(* Logix 5000 project; controller _GigaDiscovery vendor 1 type 14 code 244 rev 35.11; software revision 35.03; part 5 of 23 *)
(* tags used below, declared in another part *)
   All_RESTRAINTS_Opened : BOOL;
   Analog_Input_Pos_6 : REAL[8];
   Compressor_Pressure_OK : BOOL;
   Emergencies_CL1 : DINT[14];
   Gates_Open_Permissive : Permissive;
   Girella_Field_Actuate_During_Inactivity : BOOL;
   Girella_Gradi_Sec : DINT;
   Gondola_Axe : Axe;
   HMI_Light_Pb : BOOL;
   HMI_Status_Safety : Status_Safety;
   I_ADSL_Fault_Ch1 : BOOL;   // Gondola Communication Modem Fault CH1 -T27002C
   I_ADSL_Fault_Ch2 : BOOL;   // Gondola Communication Modem Fault CH2 -T27002C
   I_Compressor_Motor_Protection : BOOL;   // Compressor Motor Protection Feedback -F18002C
   I_Dryer_Motor_Protection : BOOL;   // Dryer Motor Protection Feedback -F18202C
   I_Gate_1_Opened : BOOL;   // Gate 1 RFID Sensor Closed -B24501J
   I_Gate_2_Opened : BOOL;   // Gate 2 RFID Sensor Closed -B24601J
   I_Gate_3_Opened : BOOL;   // Gate 3 RFID Sensor Closed -B24701J
   I_Gate_4_Opened : BOOL;   // Gate 4 RFID Sensor Closed -B24801J
   I_Light_Selector : BOOL;   // Light Selector Switch -S30408F
   I_Motor_1_2_Fan_Protection_Feedback : BOOL;   // Motor 1-2 Fan Protection Feedback -F10402C -F10406C
   I_Motor_1_Overvoltage_Control : BOOL;   // Motor 1 Overvoltage control - Relay OK -K10302G
   I_Motor_1_Thermal_Probe : BOOL;   // Motor 1 Thermal Probe -K10702H
   I_Motor_2_Overvoltage_Control : BOOL;   // Motor 2 Overvoltage control - Relay OK -K10307G
   I_Motor_2_Thermal_Probe : BOOL;   // Motor 2 Thermal Probe -K10704H
   I_Motor_3_4_Fan_Protection_Feedback : BOOL;   // Motor 3-4 Fan Protection Feedback -F12402C -F12406C
   I_Motor_3_Overvoltage_Control : BOOL;   // Motor 3 Overvoltage control - Relay OK -K12302G
   I_Motor_3_Thermal_Probe : BOOL;   // Motor 3 Thermal Probe -K12702H
   I_Motor_4_Overvoltage_Control : BOOL;   // Motor 4 Overvoltage control - Relay OK -K12307G
   I_Motor_4_Thermal_Probe : BOOL;   // Motor 4 Thermal Probe -K12704H
   I_Motor_5_6_Fan_Protection_Feedback : BOOL;   // Motor 5-6 Fan Protection Feedback -F14402C -F14406C
   I_Motor_5_Overvoltage_Control : BOOL;   // Motor 5 Overvoltage control - Relay OK -K14302G
   I_Motor_5_Thermal_Probe : BOOL;   // Motor 5 Thermal Probe -K14702H
   I_Motor_6_Overvoltage_Control : BOOL;   // Motor 6 Overvoltage control - Relay OK -K14307G
   I_Motor_6_Thermal_Probe : BOOL;   // Motor 6 Thermal Probe -K14704H
   I_Motor_7_Fan_Protection_Feedback : BOOL;   // Motor 7 Fan Protection Feedback -F16402C
   I_Motor_7_Thermal_Probe : BOOL;   // Motor 7 Thermal Probe -K16602H
   I_OCC_Operator_Enable_Key : BOOL;   // OCC Console Enabled -S30305F
   I_Platform_Closed : UDT_DCM;   // Platform Closed RFID Series -B22501J... -B22807J -B22801B
   I_Platform_Opened : UDT_DCM;   // Platform Opened RFID Series -Q23801J -Q23807J
   I_Remote_Connection_Enabled : BOOL;   // Remote Connection active ROUTER eWON K74A04E
   K_Speed : REAL;
   MCC_71_03 : BOOL[32];
   MODE : BOOL;   // MODE 0 = AUTO 1 = MANUAL -S30801F
   NO_SFTY_GateClosedSeries : BOOL;   // All Gates Closed and Locked
   O_Close_Gates : BOOL;
   ONP : DINT;   // Optional Not Present
   Pb_Platform_Stop : BOOL;   // Platform Stop Command -S30608F
   Platform_Close_Cycle : Sequencer;
   Platform_Close_Permissive : Permissive;
   Platform_Open_Cycle : Sequencer;
   Platform_Open_Permissive : Permissive;
   Pylon_Axe : Axe;
   Pylon_Field_Actuate_During_Inactivity : BOOL;
   Real : REAL[32];
   RESTRAINTS_Closed : BOOL;   // All RESTRAINTS Closed
   Restraints_Cycle : Sequencer;
   Restraints_Permissive : Permissive;
   Start_Permissive : Permissive;
   Start_Permissive2 : Permissive;
   Start_Stop_Cycle : Sequencer;
   Test : DCI_STOP_TEST;
   To_Sfty : Std_to_Sfty;
(* General, continued *)

ROUTINE Main   (* ladder *)
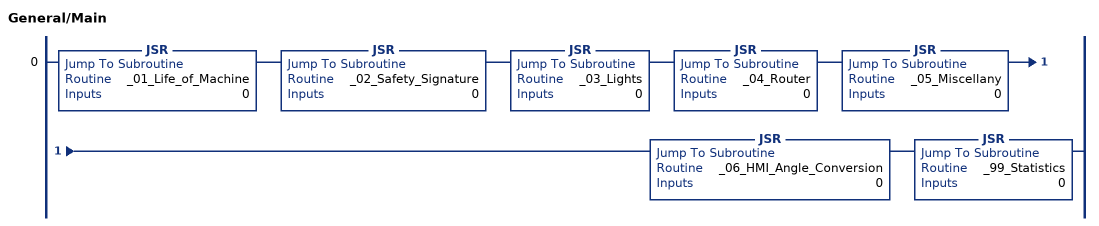
   0: JSR(_01_Life_of_Machine,0)JSR(_02_Safety_Signature,0)JSR(_03_Lights,0)JSR(_04_Router,0)JSR(_05_Miscellany,0)JSR(_06_HMI_Angle_Conversion,0)JSR(_99_Statistics,0);
END_ROUTINE
END_PROGRAM

PROGRAM HMI   (* main routine Main *)
VAR
   HMI_Auto_Cycle_Permissive : Permissive_Description := (Visible_Bits := 2147475455, Header_Description_en := 'Start Permissives (1)', Header_Description_others := 'Permessi di Start (1)', Bit_Description_en[0] := 'OCC2 Allow Main Confirm -S28602F', Bit_Description_en[1] := 'OCC Console Enabled -S30305F', Bit_Description_en[2] := 'OCC Stop Button Not Pressed -S30308F', Bit_Description_en[3] := 'All Restraints Closed', Bit_Description_en[4] := 'Gates 01-04 Closed -B24602J....-B24802J', Bit_Description_en[5] := 'Platform Stop Command Not Pressed -S30608F', Bit_Description_en[6] := 'No Emergencies Class 0', Bit_Description_en[7] := 'Restraints Proof Test Ok', Bit_Description_en[8] := 'OCC Motion Lockout -Q31203E', Bit_Description_en[9] := 'Restraints Main Valve Limit Switch Closed -B40508I', Bit_Description_en[10] := 'OCC2 E-Stop PB Not Pressed -S28502F', Bit_Description_en[11] := 'Platform Main Valve Closed -B21902I', Bit_Description_en[12] := 'Pylon Minimum Speed', Bit_Description_en[13] := 'Restraints Main Valve Pressure Switch Closed -S40602J', Bit_Description_en[14] := 'Power On Delay (80 sec.)', Bit_Description_en[15] := 'Restraints Opened Correctly', Bit_Description_en[16] := 'Restraints Pressure Switches Working Correctly', Bit_Description_en[17] := 'No Emergencies Class 1', Bit_Description_en[18] := 'Restraints Closed Correctly', Bit_Description_en[19] := 'OCC Footpedal Memory -S30901F', Bit_Description_en[20] := 'Valves Proof Test OK', Bit_Description_en[21] := 'Pylon Motors Fan On -Q9302F', Bit_Description_en[22] := 'OCC E-Stop PB Test Ok -S30301F', Bit_Description_en[23] := 'Motor Field Contactors All Disabled -Q10101E -Q10103E -Q16105E -Q16107E', Bit_Description_en[24] := 'Pylon Stopped at Home Position -B26002I -B26007I', Bit_Description_en[25] := 'Line Minimum Pressure -S21504B', Bit_Description_en[26] := 'Restraints Racks Unlock Valve Pressure Ok', Bit_Description_en[27] := 'All Racks Closed', Bit_Description_en[28] := 'Platform Opened -Q28301J -Q23807J', Bit_Description_en[29] := 'Gate Exit (G05) Closed -B25304I', Bit_Description_en[30] := 'Gate Enter (G01) Closed -B25204I', Bit_Description_en[31] := 'Gate 4 Operator(MOP) Closed -B25404J');
   HMI_Auto_Cycle_Permissive2 : Permissive_Description := (Visible_Bits := 255, Header_Description_en := 'Start Permissives (2)', Header_Description_others := 'Permessi di Start (2)', Bit_Description_en[0] := 'Platform Line Minimum Pressure Switch Closed -S21511B', Bit_Description_en[1] := 'Platform Pilot Valves Not Enabled to Open/Close -Y22002A', Bit_Description_en[2] := 'Restraints Main Valve Limit Switch Closed -B5408I', Bit_Description_en[3] := 'Restraints Sectors Left and Right Valves Unlock Disabled', Bit_Description_en[4] := 'All Restraints Sectors Disabled', Bit_Description_en[5] := 'OCC2 Stop PB Not Pressed -S28606F', Bit_Description_en[6] := 'Main Valve Closed -B40501I', Bit_Description_en[7] := 'All Restraints Sectors Racks On');
   HMI_Gates_Open_Permissive : Permissive_Description := (FailBitsConditions := 16, Visible_Bits := 190, Header_Description_en := 'Gates Open Permissives', Header_Description_others := 'Permessi di Apertura dei Cancelli', Bit_Description_en[1] := 'Ride Not in Start', Bit_Description_en[2] := 'Gondola Minimum Speed', Bit_Description_en[3] := 'Platform Main Valve Not Commanded -B21920I', Bit_Description_en[4] := 'Platform Closed -B22501J...-B22807J -B22801B', Bit_Description_en[5] := 'Pylon Safety Angle', Bit_Description_en[7] := 'Pylon Minimum Speed');
   HMI_Night_Mode : BOOL;
   HMI_Platform_Close_Error : BOOL;
   HMI_Platform_Close_Permissive : Permissive_Description := (OS_Fail := 1, Visible_Bits := 16375, Header_Description_en := 'Platform Close Permissives', Header_Description_others := 'Permessi di Chiusura della Piattaforma', Bit_Description_en[0] := 'OCC E-Stop PB Not Pressed -S30301F', Bit_Description_en[1] := 'Power On Delay (80 sec.)', Bit_Description_en[2] := 'OCC Console Enabled -S30305F', Bit_Description_en[4] := 'Motor Field Contactors All Disabled -Q10101E -Q10103E -Q16105E -Q16107E', Bit_Description_en[5] := 'Pylon Stoped At Home Position -B26002I -B26007I', Bit_Description_en[6] := 'Compressor Minimum Pressure -S21504B', Bit_Description_en[7] := 'Platform Close Alarms Not Present', Bit_Description_en[8] := 'Pylon Safety Angle', Bit_Description_en[9] := 'Pylon Minimum Speed', Bit_Description_en[10] := 'Gondola Minimun Speed', Bit_Description_en[11] := 'Platform Stop Push Button Not Pressed -S30608F', Bit_Description_en[12] := 'OCC Motion Lockout -Q31203E', Bit_Description_en[13] := 'OCC2 E-Stop PB Not Pressed -S28502F');
   HMI_Platform_Closed : BOOL := 1;
   HMI_Platform_Closing : BOOL;
   HMI_Platform_Open_Error : BOOL;
   HMI_Platform_Open_Permissive : Permissive_Description := (Visible_Bits := -2097153, Header_Description_en := 'Platform Open Permissives', Header_Description_others := 'Permessi di Apertura della Piattaforma', Bit_Description_en[0] := 'OCC E-Stop PB Not Pressed -S30301F', Bit_Description_en[1] := 'Power On Delay (80 sec.)', Bit_Description_en[2] := 'OCC Console Enabled -S3201E', Bit_Description_en[3] := 'Restraints Closed', Bit_Description_en[4] := 'Main Valve Closed -B40501I', Bit_Description_en[5] := 'Ride Not in Start', Bit_Description_en[6] := 'Compressor Minimum Pressure ', Bit_Description_en[7] := 'OCC Stop Button Not Pressed -S30308F', Bit_Description_en[8] := 'Gates 01-04 Closed -B24602J....-B24802J', Bit_Description_en[9] := 'Platform Stop Push Button not Pressed -S30608F', Bit_Description_en[10] := 'No Emergencies', Bit_Description_en[11] := 'OCC2 Allow Main Confirm -S28602F', Bit_Description_en[12] := 'OCC2 E-Stop PB Not Pressed -S28502F', Bit_Description_en[13] := 'OCC Motion Lockout -Q31203E', Bit_Description_en[14] := 'All Restraints Sectors Disabled', Bit_Description_en[15] := 'Gate Exit (G05) Closed -B25304I', Bit_Description_en[16] := 'Gate Enter (G01) Closed -B25204I', Bit_Description_en[17] := 'Gate 4 Operator(MOP) Closed -B25404J', Bit_Description_en[18] := 'Restraints Proof Test Ok', Bit_Description_en[19] := 'Restraints Main Valve Limit Switch Closed -B40508I', Bit_Description_en[20] := 'Pylon Minimum Speed', Bit_Description_en[22] := 'Restraints Opened Correctly', Bit_Description_en[23] := 'Restraints Pressure Switches Working Correctly', Bit_Description_en[24] := 'Restraints Closed Correctly', Bit_Description_en[25] := 'OCC Footpedal Memory -S30901F', Bit_Description_en[26] := 'Pylon Motors Fan On -Q9302F', Bit_Description_en[27] := 'Motor Field Contactors All Disabled -Q10101E -Q10103E -Q16105E -Q16107E', Bit_Description_en[28] := 'Pylon Stopped at Home Position -B26002I -B26007I', Bit_Description_en[29] := 'All Racks Closed', Bit_Description_en[30] := 'OCC2 Stop PB Not Pressed -S28606F', Bit_Description_en[31] := 'Platform Not at Maximum Closing Pressure -S21510B');
   HMI_Platform_Opened : BOOL;
   HMI_Platform_Opening : BOOL;
   HMI_Restraints_Closed : BOOL := 1;
   HMI_Restraints_Closing : BOOL;
   HMI_Restraints_Error : BOOL;
   HMI_Restraints_Opened : BOOL;
   HMI_Restraints_Opening : BOOL;
   HMI_Restraints_Permissive : Permissive_Description := (Visible_Bits := 7274495, Header_Description_en := 'Restraints Release Permissives', Header_Description_others := 'Permessi di Rilascio dei Maniglioni', Bit_Description_en[0] := 'OCC E-Stop PB Not Pressed -S30301F', Bit_Description_en[1] := 'Power On Delay (80 sec.)', Bit_Description_en[2] := 'OCC Console Enabled -S30305F', Bit_Description_en[3] := 'Platform Closed Cycle Complete', Bit_Description_en[4] := 'Platform Not at Maximum Closing Pressure -S21510B', Bit_Description_en[5] := 'Ride Not in Start', Bit_Description_en[6] := 'Pylon Stopped at Home Position -B26002I -B26007I', Bit_Description_en[7] := 'Pylon Encoder Low Position', Bit_Description_en[8] := 'Pylon Low Speed', Bit_Description_en[9] := 'Gondola Low Speed', Bit_Description_en[10] := 'All Pylon and Gondola Drives Not Running', Bit_Description_en[11] := 'Motor Field Contactors All Disabled -Q10101E -Q10103E -Q16105E -Q16107E', Bit_Description_en[12] := 'OCC2 E-Stop PB Not Pressed -S28502F', Bit_Description_en[13] := 'OCC Motion Lockout -Q31203E', Bit_Description_en[14] := 'Retraints Not Opened During ProofTest', Bit_Description_en[15] := 'Platform Main Valve Open -B21902I', Bit_Description_en[17] := 'Platform Line Minimum Pressure Switch Closed -S21511B', Bit_Description_en[18] := 'Platform Pilot Valves Not Enabled to Open/Close -Y22002A', Bit_Description_en[19] := 'Unlock Platform Line Pressure Switch Open -S22006B', Bit_Description_en[21] := 'Platform Closed', Bit_Description_en[22] := 'Platform Not Open');
   Os : SINT := 20;
END_VAR

ROUTINE HMI_Permissive   (* ladder *)
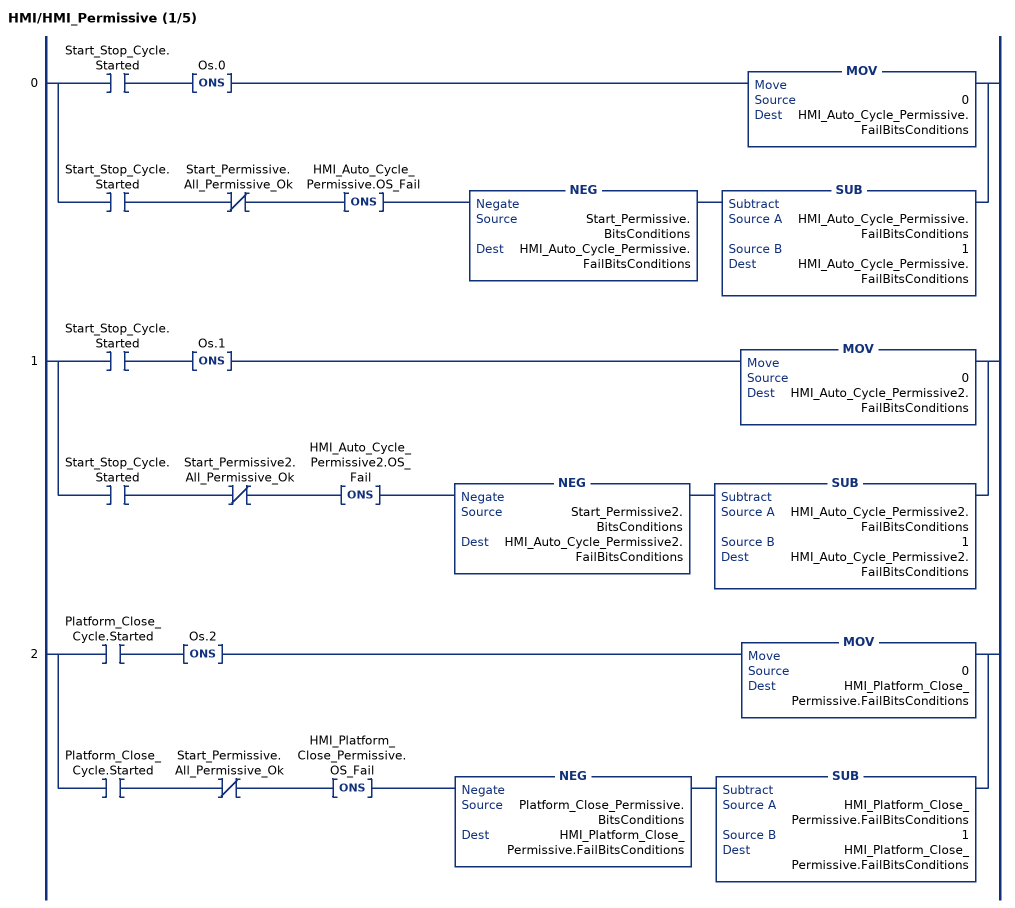
   0: [XIC(Start_Stop_Cycle.Started) ONS(Os.0) MOV(0,HMI_Auto_Cycle_Permissive.FailBitsConditions) ,XIC(Start_Stop_Cycle.Started) XIO(Start_Permissive.All_Permissive_Ok) ONS(HMI_Auto_Cycle_Permissive.OS_Fail) NEG(Start_Permissive.BitsConditions,HMI_Auto_Cycle_Permissive.FailBitsConditions) SUB(HMI_Auto_Cycle_Permissive.FailBitsConditions,1,HMI_Auto_Cycle_Permissive.FailBitsConditions) ];
   1: [XIC(Start_Stop_Cycle.Started) ONS(Os.1) MOV(0,HMI_Auto_Cycle_Permissive2.FailBitsConditions) ,XIC(Start_Stop_Cycle.Started) XIO(Start_Permissive2.All_Permissive_Ok) ONS(HMI_Auto_Cycle_Permissive2.OS_Fail) NEG(Start_Permissive2.BitsConditions,HMI_Auto_Cycle_Permissive2.FailBitsConditions) SUB(HMI_Auto_Cycle_Permissive2.FailBitsConditions,1,HMI_Auto_Cycle_Permissive2.FailBitsConditions) ];
   2: [XIC(Platform_Close_Cycle.Started) ONS(Os.2) MOV(0,HMI_Platform_Close_Permissive.FailBitsConditions) ,XIC(Platform_Close_Cycle.Started) XIO(Start_Permissive.All_Permissive_Ok) ONS(HMI_Platform_Close_Permissive.OS_Fail) NEG(Platform_Close_Permissive.BitsConditions,HMI_Platform_Close_Permissive.FailBitsConditions) SUB(HMI_Platform_Close_Permissive.FailBitsConditions,1,HMI_Platform_Close_Permissive.FailBitsConditions) ];
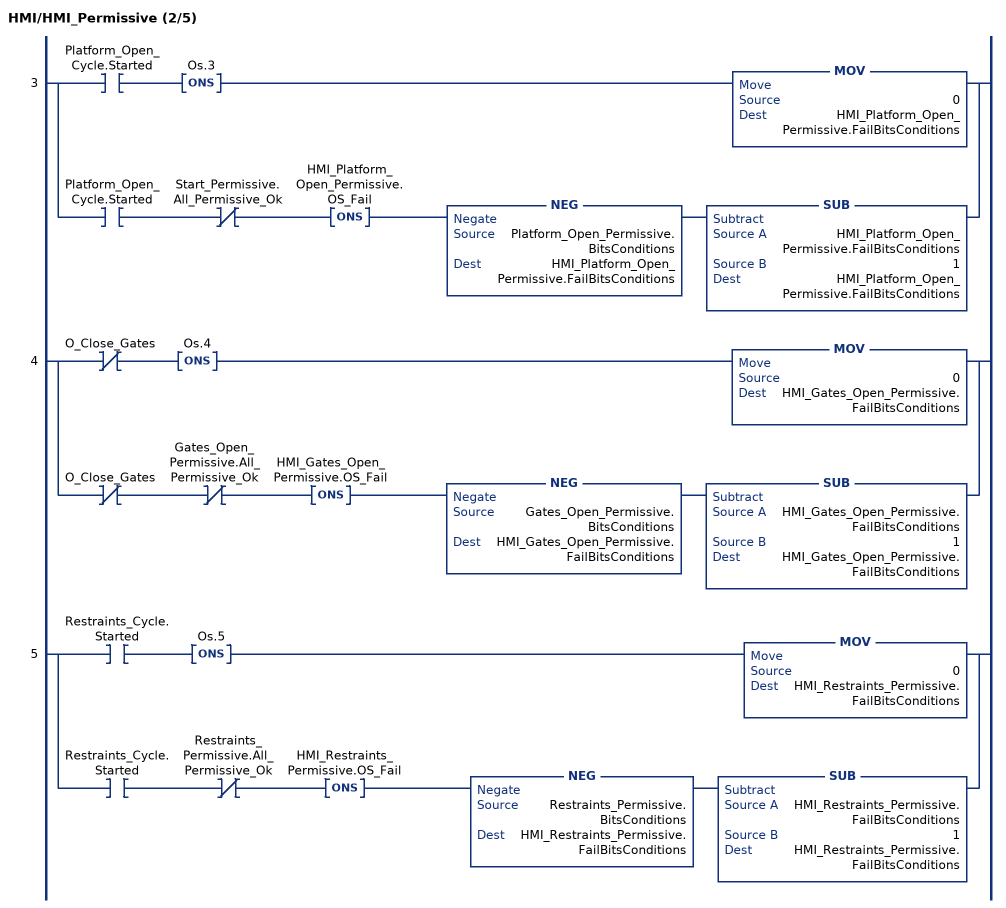
   3: [XIC(Platform_Open_Cycle.Started) ONS(Os.3) MOV(0,HMI_Platform_Open_Permissive.FailBitsConditions) ,XIC(Platform_Open_Cycle.Started) XIO(Start_Permissive.All_Permissive_Ok) ONS(HMI_Platform_Open_Permissive.OS_Fail) NEG(Platform_Open_Permissive.BitsConditions,HMI_Platform_Open_Permissive.FailBitsConditions) SUB(HMI_Platform_Open_Permissive.FailBitsConditions,1,HMI_Platform_Open_Permissive.FailBitsConditions) ];
   4: [XIO(O_Close_Gates) ONS(Os.4) MOV(0,HMI_Gates_Open_Permissive.FailBitsConditions) ,XIO(O_Close_Gates) XIO(Gates_Open_Permissive.All_Permissive_Ok) ONS(HMI_Gates_Open_Permissive.OS_Fail) NEG(Gates_Open_Permissive.BitsConditions,HMI_Gates_Open_Permissive.FailBitsConditions) SUB(HMI_Gates_Open_Permissive.FailBitsConditions,1,HMI_Gates_Open_Permissive.FailBitsConditions) ];
   5: [XIC(Restraints_Cycle.Started) ONS(Os.5) MOV(0,HMI_Restraints_Permissive.FailBitsConditions) ,XIC(Restraints_Cycle.Started) XIO(Restraints_Permissive.All_Permissive_Ok) ONS(HMI_Restraints_Permissive.OS_Fail) NEG(Restraints_Permissive.BitsConditions,HMI_Restraints_Permissive.FailBitsConditions) SUB(HMI_Restraints_Permissive.FailBitsConditions,1,HMI_Restraints_Permissive.FailBitsConditions) ];
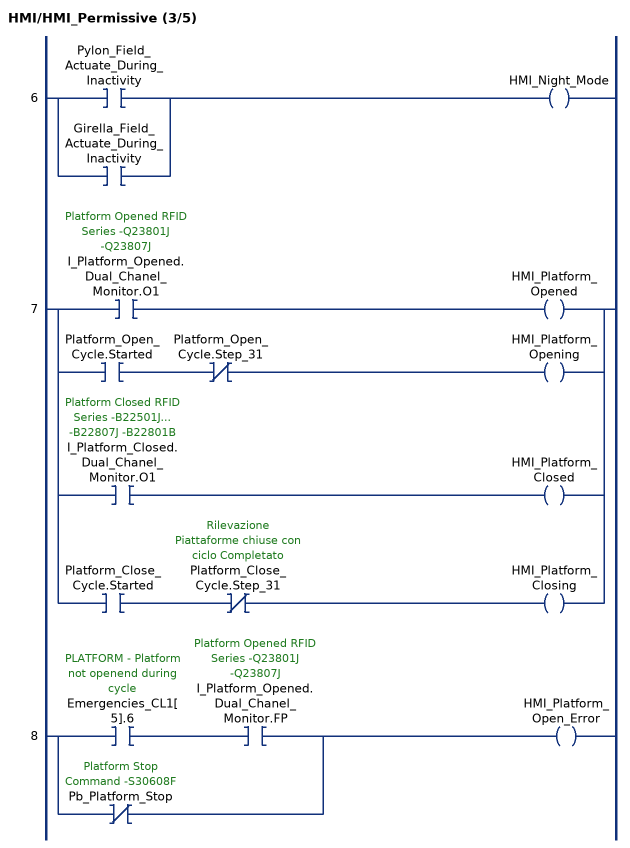
   6: [XIC(Pylon_Field_Actuate_During_Inactivity) ,XIC(Girella_Field_Actuate_During_Inactivity) ]OTE(HMI_Night_Mode);
   7: [XIC(I_Platform_Opened.Dual_Chanel_Monitor.O1) OTE(HMI_Platform_Opened) ,XIC(Platform_Open_Cycle.Started) XIO(Platform_Open_Cycle.Step_31) OTE(HMI_Platform_Opening) ,XIC(I_Platform_Closed.Dual_Chanel_Monitor.O1) OTE(HMI_Platform_Closed) ,XIC(Platform_Close_Cycle.Started) XIO(Platform_Close_Cycle.Step_31) OTE(HMI_Platform_Closing) ];
   8: [XIC(Emergencies_CL1[5].6) XIC(I_Platform_Opened.Dual_Chanel_Monitor.FP) ,XIO(Pb_Platform_Stop) ]OTE(HMI_Platform_Open_Error);
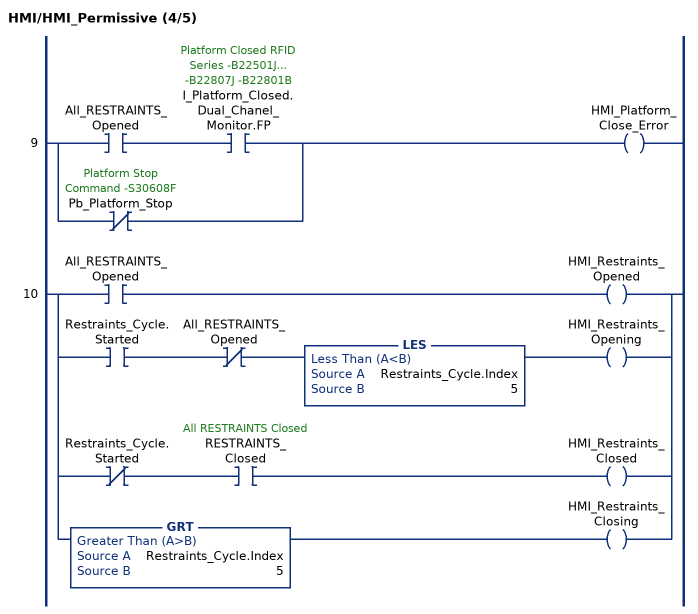
   9: [XIC(All_RESTRAINTS_Opened) XIC(I_Platform_Closed.Dual_Chanel_Monitor.FP) ,XIO(Pb_Platform_Stop) ]OTE(HMI_Platform_Close_Error);
   10: [XIC(All_RESTRAINTS_Opened) OTE(HMI_Restraints_Opened) ,XIC(Restraints_Cycle.Started) XIO(All_RESTRAINTS_Opened) LES(Restraints_Cycle.Index,5) OTE(HMI_Restraints_Opening) ,XIO(Restraints_Cycle.Started) XIC(RESTRAINTS_Closed) OTE(HMI_Restraints_Closed) ,GRT(Restraints_Cycle.Index,5) OTE(HMI_Restraints_Closing) ];
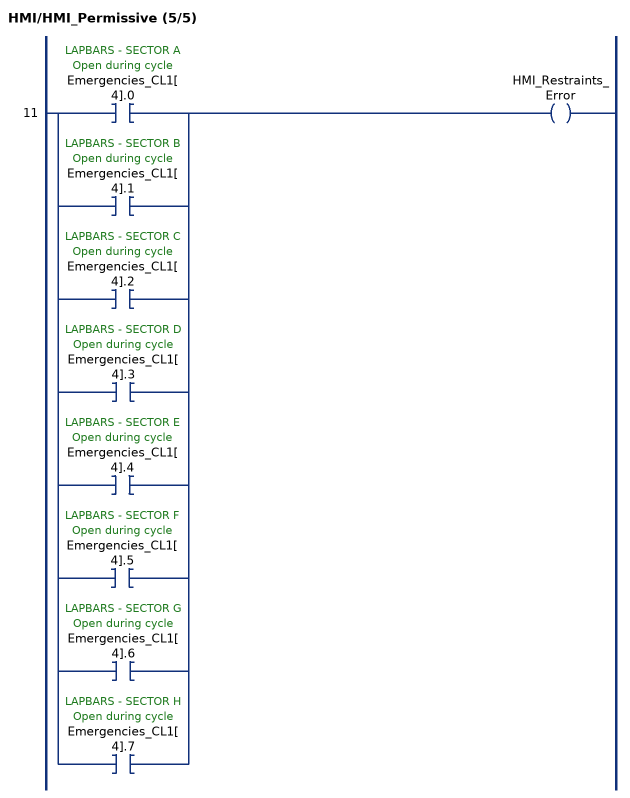
   11: [XIC(Emergencies_CL1[4].0) ,XIC(Emergencies_CL1[4].1) ,XIC(Emergencies_CL1[4].2) ,XIC(Emergencies_CL1[4].3) ,XIC(Emergencies_CL1[4].4) ,XIC(Emergencies_CL1[4].5) ,XIC(Emergencies_CL1[4].6) ,XIC(Emergencies_CL1[4].7) ]OTE(HMI_Restraints_Error);
END_ROUTINE

ROUTINE Main   (* ladder *)
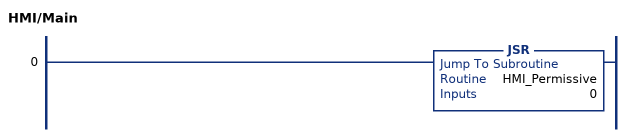
   0: JSR(HMI_Permissive,0);
END_ROUTINE
END_PROGRAM

PROGRAM Input   (* main routine Main *)
VAR
   ADD_02 : FBD_MATH := (SourceA := -11.0, SourceB := 11.0);
   ADD_03 : FBD_MATH := (SourceA := -11.0, SourceB := 11.0);
   DIV_01 : FBD_MATH := (SourceB := 100.0);
   DIV_02 : FBD_MATH := (SourceB := 100.0);
   Echo_Lights_Cmd : BOOL := 1;
   Encoder_Pulses : DINT := 4096;
   Gradi_Sec : REAL := 100.0;
   In_FGEN_01 : FUNCTION_GENERATOR := (XY1Size := 2, Out := 0.0061035156);
   In_FGEN_02 : FUNCTION_GENERATOR := (XY1Size := 2);
   In_FGEN_03 : FUNCTION_GENERATOR := (In := -2.125, XY1Size := 2, Out := -0.025939941);
   In_FGEN_04 : FUNCTION_GENERATOR := (XY1Size := 2);
   In_FGEN_05 : FUNCTION_GENERATOR := (In := -2.0625, XY1Size := 2, Out := -0.025177002);
   In_FGEN_06 : FUNCTION_GENERATOR := (XY1Size := 2);
   In_FGEN_07 : FUNCTION_GENERATOR := (In := -2.25, XY1Size := 2, Out := -0.02746582);
   In_FGEN_08 : FUNCTION_GENERATOR := (XY1Size := 2);
   In_FGEN_09 : FUNCTION_GENERATOR := (XY1Size := 2, Out := 0.0061035156);
   In_FGEN_10 : FUNCTION_GENERATOR := (XY1Size := 2);
   In_FGEN_11 : FUNCTION_GENERATOR := (In := -2.125, XY1Size := 2, Out := -0.025939941);
   In_FGEN_12 : FUNCTION_GENERATOR := (XY1Size := 2);
   In_FGEN_13 : FUNCTION_GENERATOR := (In := -2.125, XY1Size := 2, Out := -0.025939941);
   In_FGEN_14 : FUNCTION_GENERATOR := (XY1Size := 2);
   In_FGEN_15 : FUNCTION_GENERATOR := (In := -2.375, XY1Size := 2, Out := -0.0289917);
   In_FGEN_16 : FUNCTION_GENERATOR := (XY1Size := 2);
   Input_Scalaggi : Scale_2_P[16] := ([0].Input[1] := 10.0, [0].Output[1] := 10000.0, [1].Input[1] := 10.0, [1].Output[1] := 10000.0, [2].Input[1] := 10.0, [2].Output[1] := 10000.0, [3].Input[1] := 10.0, [3].Output[1] := 10000.0, [4].Input[0] := -32768.0, [4].Input[1] := 32767.0, [4].Output[0] := -400.0, [4].Output[1] := 400.0, [5].Input[0] := -32767.0, [5].Input[1] := 32767.0, [5].Output[0] := -500.0, [5].Output[1] := 500.0, [6].Input[0] := -32767.0, [6].Input[1] := 32767.0, [6].Output[0] := -400.0, [6].Output[1] := 400.0, [7].Input[0] := -32767.0, [7].Input[1] := 32767.0, [7].Output[0] := -500.0, [7].Output[1] := 500.0, [8].Input[0] := -32767.0, [8].Input[1] := 32767.0, [8].Output[0] := -400.0, [8].Output[1] := 400.0, [9].Input[0] := -32767.0, [9].Input[1] := 32767.0, [9].Output[0] := -100.0, [9].Output[1] := 100.0, [10].Input[0] := -32767.0, [10].Input[1] := 32767.0, [10].Output[0] := -400.0, [10].Output[1] := 400.0, [11].Input[0] := -32767.0, [11].Input[1] := 32767.0, [11].Output[0] := -500.0, [11].Output[1] := 500.0);
   Lights_Cmd : BOOL := 1;
   LPF_01 : FILTER_LOW_PASS := (WLag := 1.7453293, Order := 1, RTSTime := 1, DeltaT := 0.001);
   LPF_02 : FILTER_LOW_PASS := (WLag := 0.34906584, Order := 1, RTSTime := 1, DeltaT := 0.001);
   LPF_03 : FILTER_LOW_PASS := (WLag := 1.7453293, Order := 1, RTSTime := 1, DeltaT := 0.001);
   LPF_04 : FILTER_LOW_PASS := (In := -0.025939941, Order := 1, RTSTime := 1, Out := -0.02593994, DeltaT := 0.001, Status := 16#0000_0003, InstructFault := 1, WLagInv := 1);
   LPF_05 : FILTER_LOW_PASS := (WLag := 2.0, Order := 2, RTSTime := 1, DeltaT := 0.001);
   LPF_06 : FILTER_LOW_PASS := (WLag := 0.34906584, Order := 1, RTSTime := 1, Out := -2.877214e-24, DeltaT := 0.001);
   LPF_07 : FILTER_LOW_PASS := (In := -0.025939941, Order := 1, RTSTime := 1, Out := -0.025939941, DeltaT := 0.001, Status := 16#0000_0003, InstructFault := 1, WLagInv := 1);
   LPF_08 : FILTER_LOW_PASS := (WLag := 2.0, Order := 2, RTSTime := 1, DeltaT := 0.001);
   Os : DINT;
        .0   // USED
   Pignone : DINT := 20;
   Pylon_Axe_Position_360_SUB : REAL := -1487274.9;
   RAD_01 : FBD_MATH_ADVANCED := (Source := 100.0, Dest := 1.7453293);
   RAD_02 : FBD_MATH_ADVANCED := (Source := 20.0, Dest := 0.34906584);
   RAD_03 : FBD_MATH_ADVANCED := (Source := 100.0, Dest := 1.7453293);
   RAD_04 : FBD_MATH_ADVANCED := (Source := 20.0, Dest := 0.34906584);
   Ralla : DINT := 145;
   RallaPignone : REAL := 7.25;
   Riduttore : REAL := 17.5;
   Timer : TIMER[50] := ([0].PRE := 2000, [0].ACC := 2000, [0].EN := 1, [0].DN := 1, [1].PRE := 500, [2].PRE := 500, [3].PRE := 500, [4].PRE := 500, [5].PRE := 500, [6].PRE := 500, [7].PRE := 500, [8].PRE := 500, [9].PRE := 500, [10].PRE := 500, [11].PRE := 500, [12].PRE := 500, [13].PRE := 500, [14].PRE := 500, [15].PRE := 500, [16].PRE := 500, [17].PRE := 500, [18].PRE := 500, [19].PRE := 500, [20].PRE := 500, [21].PRE := 500, [22].PRE := 500, [23].PRE := 500, [24].PRE := 500, [25].PRE := 500, [26].PRE := 500, [27].PRE := 500, [28].PRE := 500, [29].PRE := 500, [30].PRE := 500, [31].PRE := 500, [32].PRE := 500, [33].PRE := 500, [34].PRE := 500, [35].PRE := 500, [36].PRE := 500, [37].PRE := 500, [38].PRE := 500, [39].PRE := 500, [40].PRE := 500, [41].PRE := 5000, [41].ACC := 5000, [41].EN := 1, [41].DN := 1, [42].PRE := 500, [49].PRE := 300000, [49].ACC := 300000, [49].EN := 1, [49].DN := 1);
   ToBe_Define_Std : DINT := 10819;
   TobeDefine_real : REAL;
END_VAR

ROUTINE _01_Input_Map_Analog   (* function block diagram *)
   SHEET 1   // Pilone
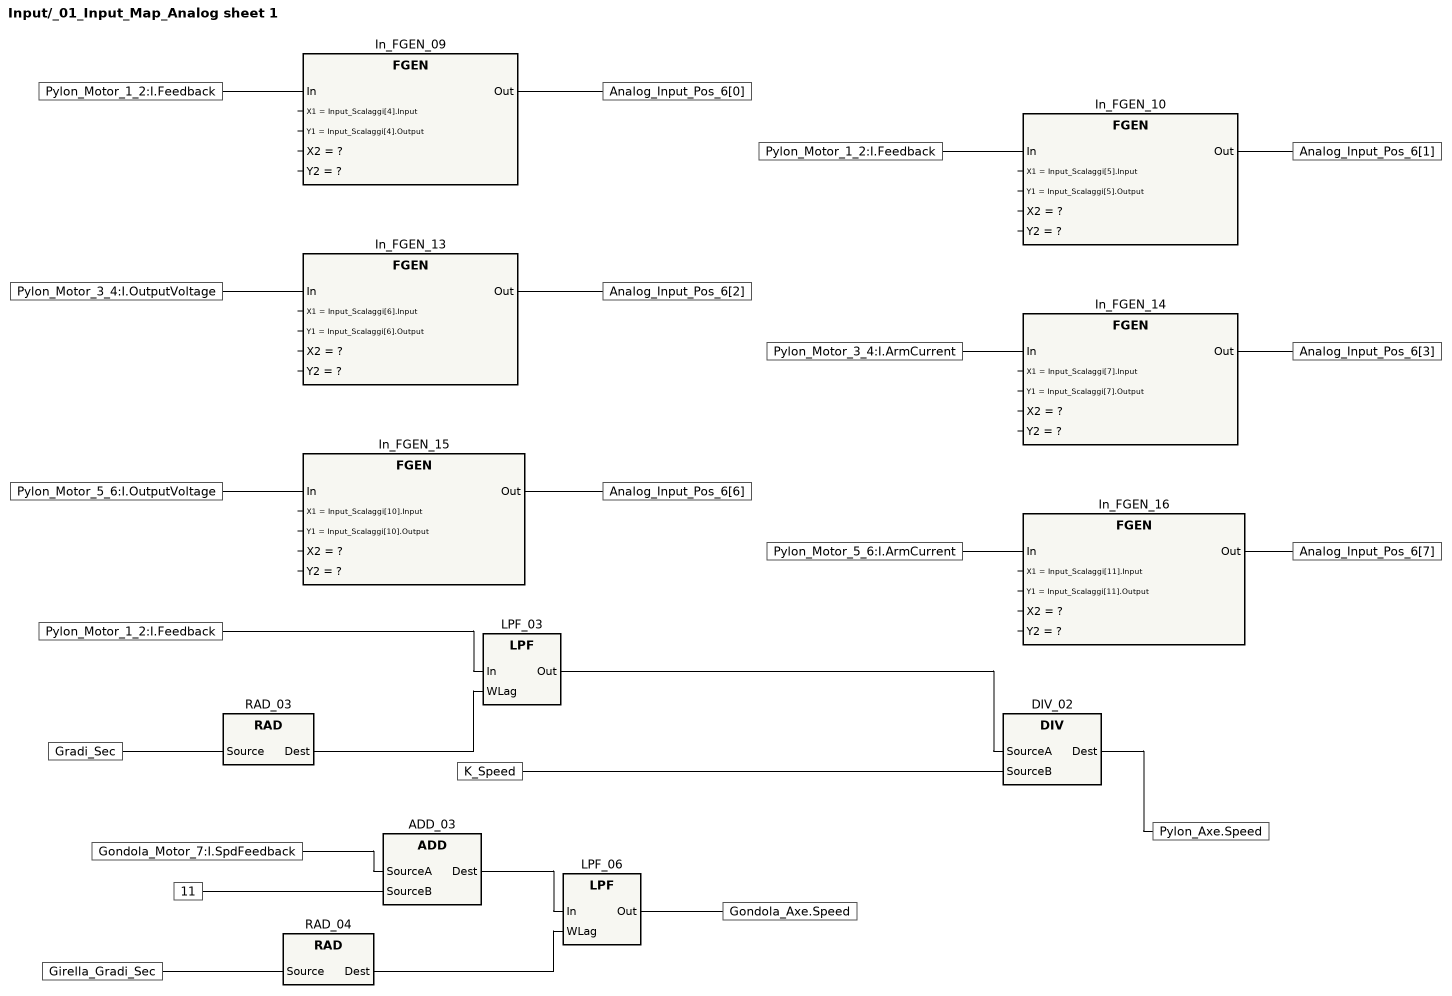
   RAD_03 : RAD(Source := Gradi_Sec);
   RAD_04 : RAD(Source := Girella_Gradi_Sec);
   In_FGEN_09 : FGEN(In := Pylon_Motor_1_2:I.Feedback, X1 := Input_Scalaggi[4].Input, Y1 := Input_Scalaggi[4].Output, X2 := ?, Y2 := ?);
   In_FGEN_13 : FGEN(In := Pylon_Motor_3_4:I.OutputVoltage, X1 := Input_Scalaggi[6].Input, Y1 := Input_Scalaggi[6].Output, X2 := ?, Y2 := ?);
   In_FGEN_15 : FGEN(In := Pylon_Motor_5_6:I.OutputVoltage, X1 := Input_Scalaggi[10].Input, Y1 := Input_Scalaggi[10].Output, X2 := ?, Y2 := ?);
   ADD_03 : ADD(SourceA := Gondola_Motor_7:I.SpdFeedback, SourceB := 11);
   LPF_03 : LPF(In := Pylon_Motor_1_2:I.Feedback, WLag := RAD_03.Dest);
   LPF_06 : LPF(In := ADD_03.Dest, WLag := RAD_04.Dest);
   Analog_Input_Pos_6[0] := In_FGEN_09.Out;
   Analog_Input_Pos_6[2] := In_FGEN_13.Out;
   Analog_Input_Pos_6[6] := In_FGEN_15.Out;
   Gondola_Axe.Speed := LPF_06.Out;
   DIV_02 : DIV(SourceA := LPF_03.Out, SourceB := K_Speed);
   In_FGEN_10 : FGEN(In := Pylon_Motor_1_2:I.Feedback, X1 := Input_Scalaggi[5].Input, Y1 := Input_Scalaggi[5].Output, X2 := ?, Y2 := ?);
   In_FGEN_14 : FGEN(In := Pylon_Motor_3_4:I.ArmCurrent, X1 := Input_Scalaggi[7].Input, Y1 := Input_Scalaggi[7].Output, X2 := ?, Y2 := ?);
   In_FGEN_16 : FGEN(In := Pylon_Motor_5_6:I.ArmCurrent, X1 := Input_Scalaggi[11].Input, Y1 := Input_Scalaggi[11].Output, X2 := ?, Y2 := ?);
   Pylon_Axe.Speed := DIV_02.Dest;
   Analog_Input_Pos_6[1] := In_FGEN_10.Out;
   Analog_Input_Pos_6[3] := In_FGEN_14.Out;
   Analog_Input_Pos_6[7] := In_FGEN_16.Out;
   SHEET 2   // Gondola
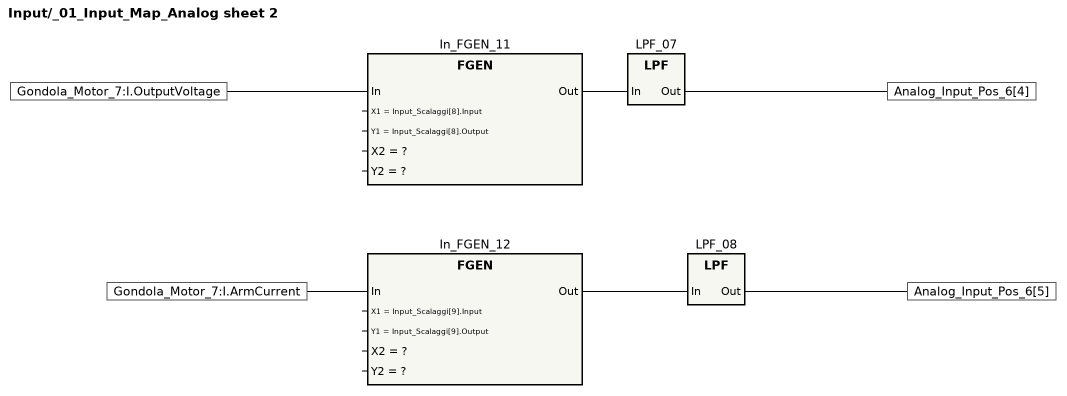
   In_FGEN_11 : FGEN(In := Gondola_Motor_7:I.OutputVoltage, X1 := Input_Scalaggi[8].Input, Y1 := Input_Scalaggi[8].Output, X2 := ?, Y2 := ?);
   In_FGEN_12 : FGEN(In := Gondola_Motor_7:I.ArmCurrent, X1 := Input_Scalaggi[9].Input, Y1 := Input_Scalaggi[9].Output, X2 := ?, Y2 := ?);
   LPF_07 : LPF(In := In_FGEN_11.Out);
   LPF_08 : LPF(In := In_FGEN_12.Out);
   Analog_Input_Pos_6[4] := LPF_07.Out;
   Analog_Input_Pos_6[5] := LPF_08.Out;
END_ROUTINE

ROUTINE _01_Primary_OCC   (* ladder *)
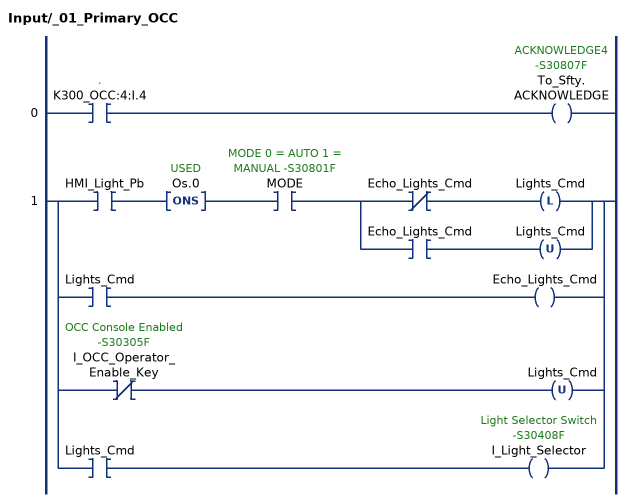
   0: XIC(K300_OCC:4:I.4)OTE(To_Sfty.ACKNOWLEDGE);
   1: [XIC(HMI_Light_Pb) ONS(Os.0) XIC(MODE) [XIO(Echo_Lights_Cmd) OTL(Lights_Cmd) ,XIC(Echo_Lights_Cmd) OTU(Lights_Cmd) ] ,XIC(Lights_Cmd) OTE(Echo_Lights_Cmd) ,XIO(I_OCC_Operator_Enable_Key) OTU(Lights_Cmd) ,XIC(Lights_Cmd) OTE(I_Light_Selector) ];
END_ROUTINE

ROUTINE _02_Secondary_OCC   (* ladder *)
END_ROUTINE

ROUTINE _03_MCC   (* ladder *)
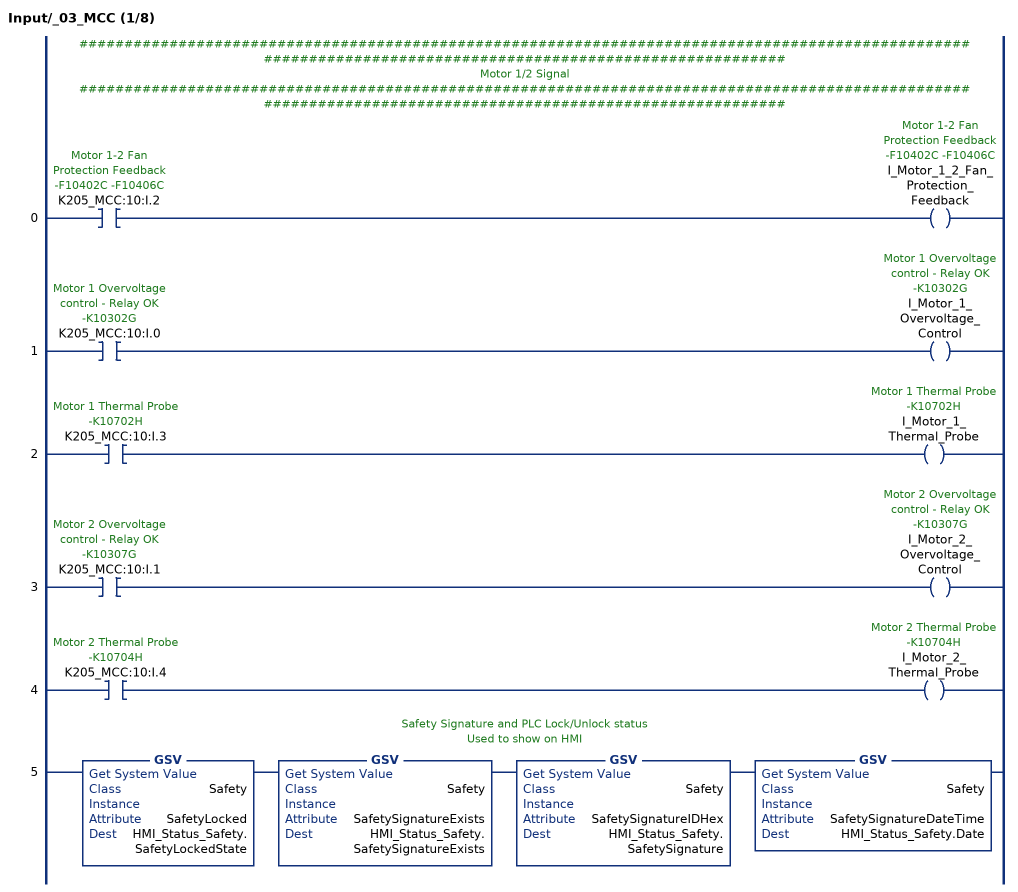
   // #############################################################################################################################################################
   // Motor 1/2 Signal
   // #############################################################################################################################################################
   0: XIC(K205_MCC:10:I.2)OTE(I_Motor_1_2_Fan_Protection_Feedback);
   1: XIC(K205_MCC:10:I.0)OTE(I_Motor_1_Overvoltage_Control);
   2: XIC(K205_MCC:10:I.3)OTE(I_Motor_1_Thermal_Probe);
   3: XIC(K205_MCC:10:I.1)OTE(I_Motor_2_Overvoltage_Control);
   4: XIC(K205_MCC:10:I.4)OTE(I_Motor_2_Thermal_Probe);
   // Safety Signature and PLC Lock/Unlock status
   // Used to show on HMI
   5: GSV(Safety,,SafetyLocked,HMI_Status_Safety.SafetyLockedState)GSV(Safety,,SafetySignatureExists,HMI_Status_Safety.SafetySignatureExists)GSV(Safety,,SafetySignatureIDHex,HMI_Status_Safety.SafetySignature)GSV(Safety,,SafetySignatureDateTime,HMI_Status_Safety.Date);
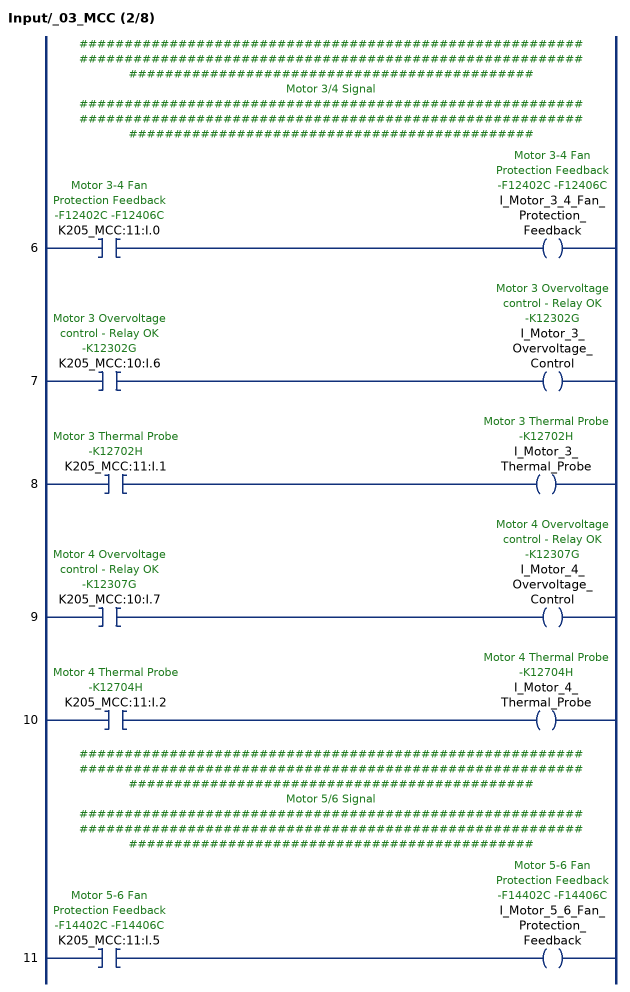
   // #############################################################################################################################################################
   // Motor 3/4 Signal
   // #############################################################################################################################################################
   6: XIC(K205_MCC:11:I.0)OTE(I_Motor_3_4_Fan_Protection_Feedback);
   7: XIC(K205_MCC:10:I.6)OTE(I_Motor_3_Overvoltage_Control);
   8: XIC(K205_MCC:11:I.1)OTE(I_Motor_3_Thermal_Probe);
   9: XIC(K205_MCC:10:I.7)OTE(I_Motor_4_Overvoltage_Control);
   10: XIC(K205_MCC:11:I.2)OTE(I_Motor_4_Thermal_Probe);
   // #############################################################################################################################################################
   // Motor 5/6 Signal
   // #############################################################################################################################################################
   11: XIC(K205_MCC:11:I.5)OTE(I_Motor_5_6_Fan_Protection_Feedback);
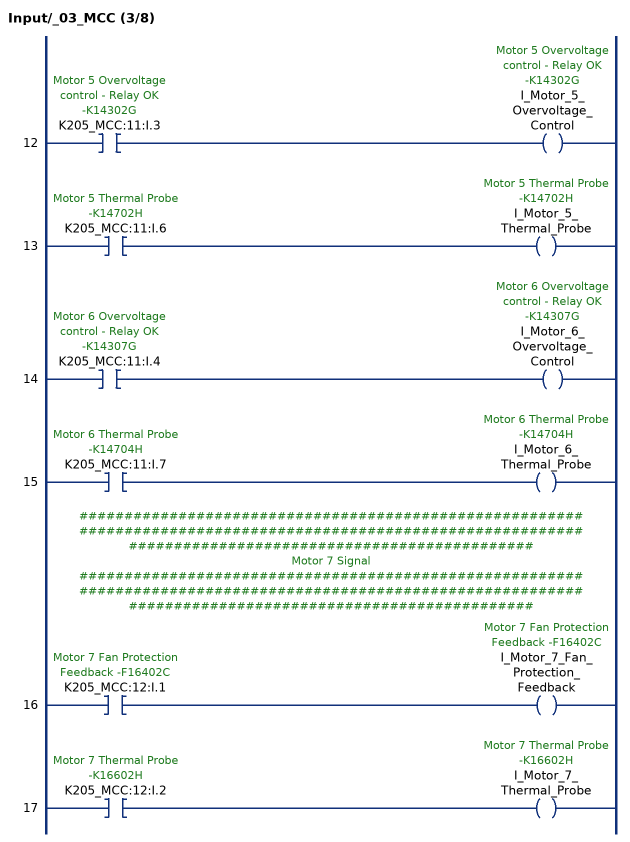
   12: XIC(K205_MCC:11:I.3)OTE(I_Motor_5_Overvoltage_Control);
   13: XIC(K205_MCC:11:I.6)OTE(I_Motor_5_Thermal_Probe);
   14: XIC(K205_MCC:11:I.4)OTE(I_Motor_6_Overvoltage_Control);
   15: XIC(K205_MCC:11:I.7)OTE(I_Motor_6_Thermal_Probe);
   // #############################################################################################################################################################
   // Motor 7 Signal
   // #############################################################################################################################################################
   16: XIC(K205_MCC:12:I.1)OTE(I_Motor_7_Fan_Protection_Feedback);
   17: XIC(K205_MCC:12:I.2)OTE(I_Motor_7_Thermal_Probe);
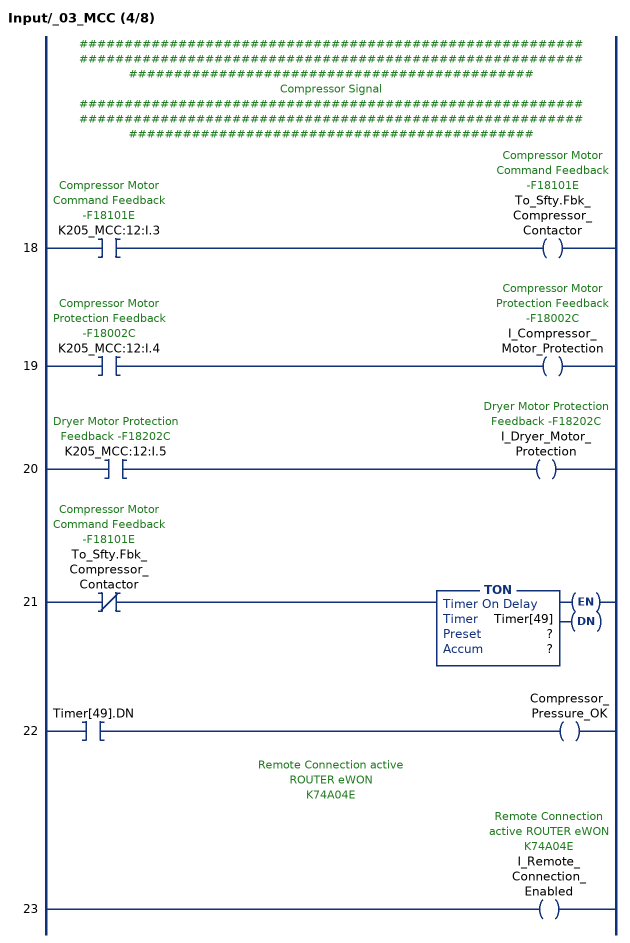
   // #############################################################################################################################################################
   // Compressor Signal
   // #############################################################################################################################################################
   18: XIC(K205_MCC:12:I.3)OTE(To_Sfty.Fbk_Compressor_Contactor);
   19: XIC(K205_MCC:12:I.4)OTE(I_Compressor_Motor_Protection);
   20: XIC(K205_MCC:12:I.5)OTE(I_Dryer_Motor_Protection);
   21: XIO(To_Sfty.Fbk_Compressor_Contactor)TON(Timer[49],?,?);
   22: XIC(Timer[49].DN)OTE(Compressor_Pressure_OK);
   // Remote Connection active
   // ROUTER eWON
   // K74A04E
   23: OTE(I_Remote_Connection_Enabled);
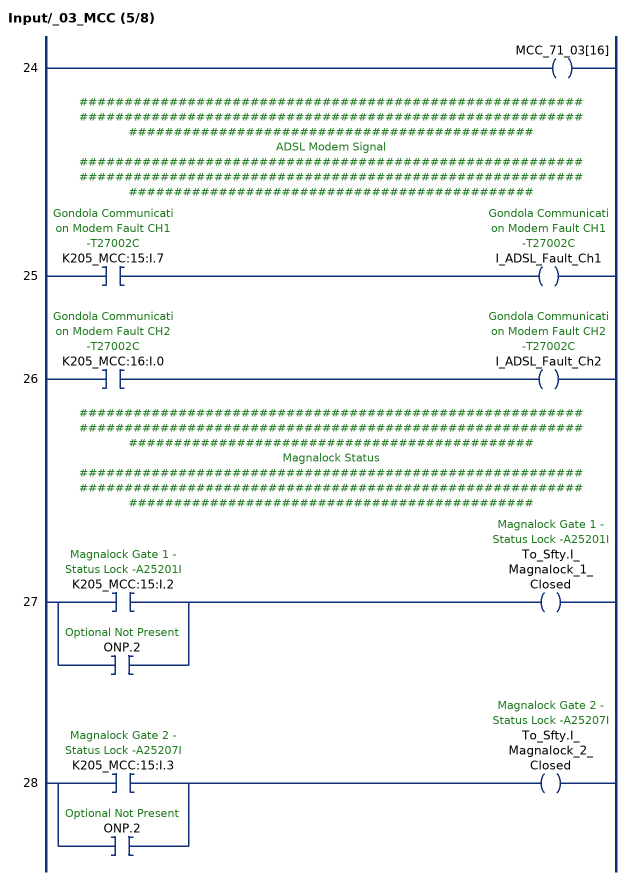
   24: OTE(MCC_71_03[16]);
   // #############################################################################################################################################################
   // ADSL Modem Signal
   // #############################################################################################################################################################
   25: XIC(K205_MCC:15:I.7)OTE(I_ADSL_Fault_Ch1);
   26: XIC(K205_MCC:16:I.0)OTE(I_ADSL_Fault_Ch2);
   // #############################################################################################################################################################
   // Magnalock Status
   // #############################################################################################################################################################
   27: [XIC(K205_MCC:15:I.2) ,XIC(ONP.2) ]OTE(To_Sfty.I_Magnalock_1_Closed);
   28: [XIC(K205_MCC:15:I.3) ,XIC(ONP.2) ]OTE(To_Sfty.I_Magnalock_2_Closed);
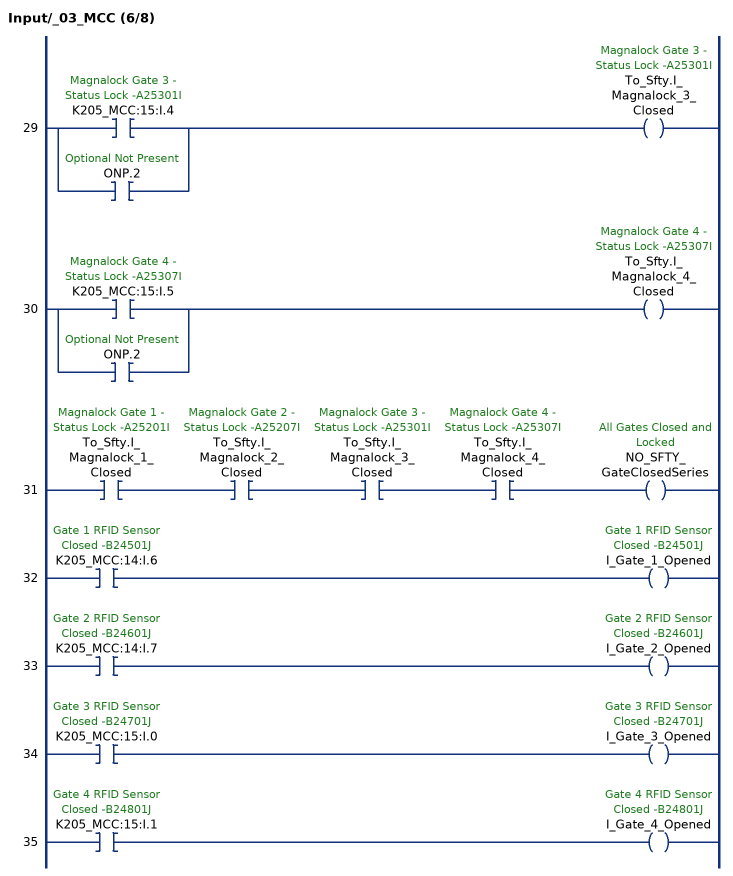
   29: [XIC(K205_MCC:15:I.4) ,XIC(ONP.2) ]OTE(To_Sfty.I_Magnalock_3_Closed);
   30: [XIC(K205_MCC:15:I.5) ,XIC(ONP.2) ]OTE(To_Sfty.I_Magnalock_4_Closed);
   31: XIC(To_Sfty.I_Magnalock_1_Closed)XIC(To_Sfty.I_Magnalock_2_Closed)XIC(To_Sfty.I_Magnalock_3_Closed)XIC(To_Sfty.I_Magnalock_4_Closed)OTE(NO_SFTY_GateClosedSeries);
   32: XIC(K205_MCC:14:I.6)OTE(I_Gate_1_Opened);
   33: XIC(K205_MCC:14:I.7)OTE(I_Gate_2_Opened);
   34: XIC(K205_MCC:15:I.0)OTE(I_Gate_3_Opened);
   35: XIC(K205_MCC:15:I.1)OTE(I_Gate_4_Opened);
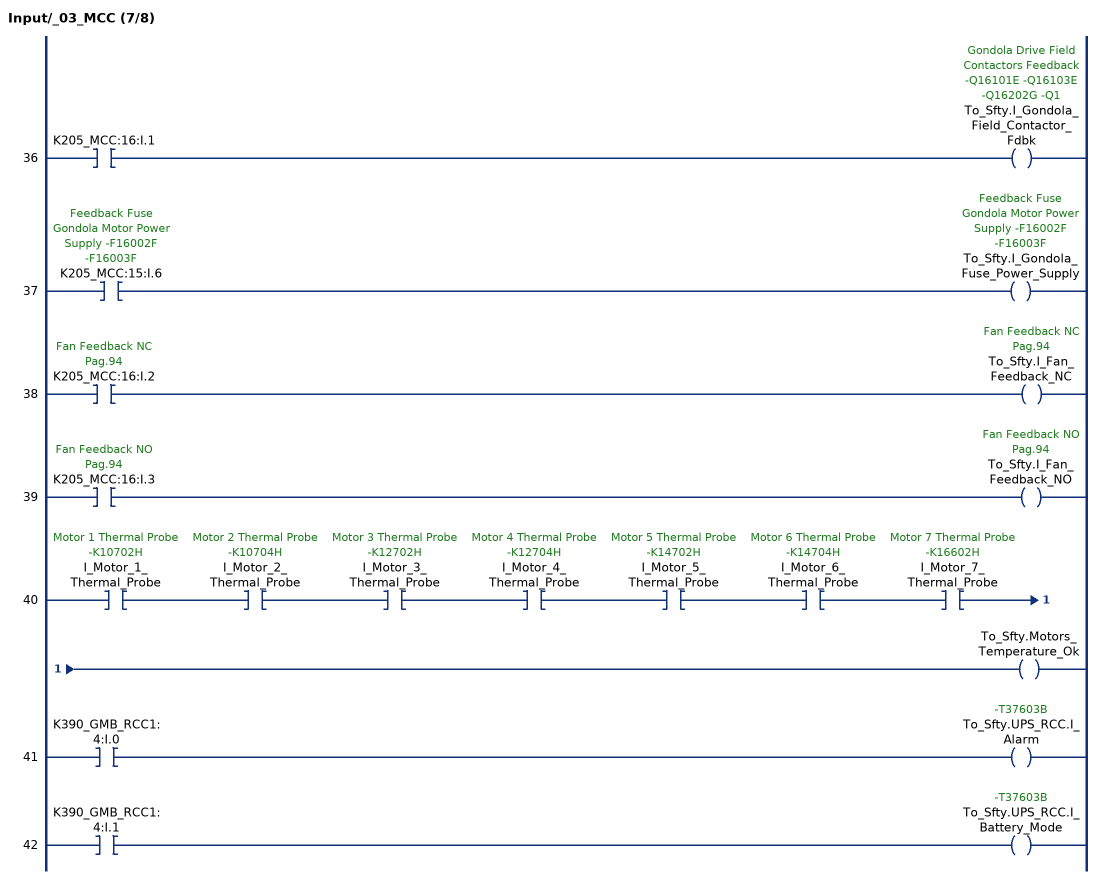
   36: XIC(K205_MCC:16:I.1)OTE(To_Sfty.I_Gondola_Field_Contactor_Fdbk);
   37: XIC(K205_MCC:15:I.6)OTE(To_Sfty.I_Gondola_Fuse_Power_Supply);
   38: XIC(K205_MCC:16:I.2)OTE(To_Sfty.I_Fan_Feedback_NC);
   39: XIC(K205_MCC:16:I.3)OTE(To_Sfty.I_Fan_Feedback_NO);
   40: XIC(I_Motor_1_Thermal_Probe)XIC(I_Motor_2_Thermal_Probe)XIC(I_Motor_3_Thermal_Probe)XIC(I_Motor_4_Thermal_Probe)XIC(I_Motor_5_Thermal_Probe)XIC(I_Motor_6_Thermal_Probe)XIC(I_Motor_7_Thermal_Probe)OTE(To_Sfty.Motors_Temperature_Ok);
   41: XIC(K390_GMB_RCC1:4:I.0)OTE(To_Sfty.UPS_RCC.I_Alarm);
   42: XIC(K390_GMB_RCC1:4:I.1)OTE(To_Sfty.UPS_RCC.I_Battery_Mode);
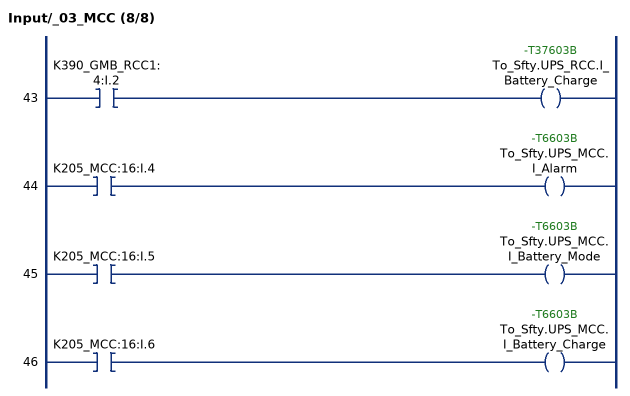
   43: XIC(K390_GMB_RCC1:4:I.2)OTE(To_Sfty.UPS_RCC.I_Battery_Charge);
   44: XIC(K205_MCC:16:I.4)OTE(To_Sfty.UPS_MCC.I_Alarm);
   45: XIC(K205_MCC:16:I.5)OTE(To_Sfty.UPS_MCC.I_Battery_Mode);
   46: XIC(K205_MCC:16:I.6)OTE(To_Sfty.UPS_MCC.I_Battery_Charge);
END_ROUTINE
